// TIA Portal project "Catalyst_syzygy_v2.1" (V17) (continued)
VERSION : 0.1
   VAR
      ConnectP : TCON_IP_v4;
      MBControl : Struct
         diconnect : Bool;
      END_STRUCT;
   END_VAR
BEGIN
   ConnectP.InterfaceId := 258;
   ConnectP.ID := 16#1;
   ConnectP.ConnectionType := 11;
   ConnectP.LocalPort := 502;
END_DATA_BLOCK

DATA_BLOCK "TC-402B_DB"   // DB425
{ S7_Optimized_Access := 'TRUE' }
VERSION : 0.1
   VAR
      Data : "EurothermCtls_UDT";
      AddrCtrl : Struct
         CurrentAddr : UDInt;
         Down : Bool;
         Up : Bool;
         RisingUp : Bool;
      END_STRUCT;
   END_VAR
BEGIN
END_DATA_BLOCK

DATA_BLOCK "TC-402B_R1"   // DB429
{ S7_Optimized_Access := 'TRUE' }
AUTHOR : JL
VERSION : 0.1
// stored: InstanceOfName Eurotherm_MB_FB
"Eurotherm_MB_FB"
BEGIN
END_DATA_BLOCK

DATA_BLOCK "TC-402B_R2"   // DB431
{ S7_Optimized_Access := 'TRUE' }
AUTHOR : JL
VERSION : 0.1
// stored: InstanceOfName Eurotherm_MB_FB
"Eurotherm_MB_FB"
BEGIN
END_DATA_BLOCK

DATA_BLOCK "TC-402B_R3"   // DB432
{ S7_Optimized_Access := 'TRUE' }
AUTHOR : JL
VERSION : 0.1
// stored: InstanceOfName Eurotherm_MB_FB
"Eurotherm_MB_FB"
BEGIN
END_DATA_BLOCK

DATA_BLOCK "TC-402B_W1"   // DB435
{ S7_Optimized_Access := 'TRUE' }
AUTHOR : JL
VERSION : 0.1
// stored: InstanceOfName Eurotherm_MB_FB
"Eurotherm_MB_FB"
BEGIN
END_DATA_BLOCK

// folder: Outside Comms/ModBus Comms/MFCs/MFC-4011

DATA_BLOCK "MFC-4011_MB_R_DB"   // DB93
{ S7_Optimized_Access := 'TRUE' }
VERSION : 0.1
// stored: InstanceOfName MFC_MB_rDT
"MFC_MB_rDT"
BEGIN
END_DATA_BLOCK

DATA_BLOCK "MFC-4011_MB_W_DB"   // DB130
{ S7_Optimized_Access := 'TRUE' }
VERSION : 0.1
// stored: InstanceOfName MFC_MB_rDT
"MFC_MB_rDT"
BEGIN
END_DATA_BLOCK

DATA_BLOCK "MFC-4011_MB_RCMD_DB"   // DB133
{ S7_Optimized_Access := 'TRUE' }
AUTHOR : JL
VERSION : 0.1
// stored: InstanceOfName MFC_MB_iDT
"MFC_MB_iDT"
BEGIN
END_DATA_BLOCK

DATA_BLOCK "MFC-4011_MB_WCMD_DB"   // DB139
{ S7_Optimized_Access := 'TRUE' }
AUTHOR : JL
VERSION : 0.1
// stored: InstanceOfName MFC_MB_iDT
"MFC_MB_iDT"
BEGIN
END_DATA_BLOCK

DATA_BLOCK "MFC-4011_DB_MB"   // DB144
TITLE = MFC-4011 Modbus DB
{ S7_Optimized_Access := 'TRUE' }
VERSION : 0.1
   VAR
      Data : "AlicatCtl_UDT";
   END_VAR
BEGIN
END_DATA_BLOCK

// folder: Outside Comms/ModBus Comms/MFCs/MFC-4012

DATA_BLOCK "MFC-4012_MB_R_DB"   // DB200
{ S7_Optimized_Access := 'TRUE' }
VERSION : 0.1
// stored: InstanceOfName MFC_MB_rDT
"MFC_MB_rDT"
BEGIN
END_DATA_BLOCK

DATA_BLOCK "MFC-4012_MB_W_DB"   // DB201
{ S7_Optimized_Access := 'TRUE' }
VERSION : 0.1
// stored: InstanceOfName MFC_MB_rDT
"MFC_MB_rDT"
BEGIN
END_DATA_BLOCK

DATA_BLOCK "MFC-4012_MB_RCMD_DB"   // DB202
{ S7_Optimized_Access := 'TRUE' }
AUTHOR : JL
VERSION : 0.1
// stored: InstanceOfName MFC_MB_iDT
"MFC_MB_iDT"
BEGIN
END_DATA_BLOCK

DATA_BLOCK "MFC-4012_MB_WCMD_DB"   // DB239
{ S7_Optimized_Access := 'TRUE' }
AUTHOR : JL
VERSION : 0.1
// stored: InstanceOfName MFC_MB_iDT
"MFC_MB_iDT"
BEGIN
END_DATA_BLOCK

DATA_BLOCK "MFC-4012_DB_MB"   // DB240
TITLE = MFC-4011 Modbus DB
{ S7_Optimized_Access := 'TRUE' }
VERSION : 0.1
   VAR
      Data : "AlicatCtl_UDT";
   END_VAR
BEGIN
END_DATA_BLOCK

// folder: Outside Comms/ModBus Comms/MFCs/MFC-4021

DATA_BLOCK "MFC-4021_MB_R_DB"   // DB421
{ S7_Optimized_Access := 'TRUE' }
VERSION : 0.1
// stored: InstanceOfName MFC_MB_rDT
"MFC_MB_rDT"
BEGIN
END_DATA_BLOCK

DATA_BLOCK "MFC-4021_MB_W_DB"   // DB422
{ S7_Optimized_Access := 'TRUE' }
VERSION : 0.1
// stored: InstanceOfName MFC_MB_rDT
"MFC_MB_rDT"
BEGIN
END_DATA_BLOCK

DATA_BLOCK "MFC-4021_MB_RCMD_DB"   // DB423
{ S7_Optimized_Access := 'TRUE' }
AUTHOR : JL
VERSION : 0.1
// stored: InstanceOfName MFC_MB_iDT
"MFC_MB_iDT"
BEGIN
END_DATA_BLOCK

DATA_BLOCK "MFC-4021_MB_WCMD_DB"   // DB426
{ S7_Optimized_Access := 'TRUE' }
AUTHOR : JL
VERSION : 0.1
// stored: InstanceOfName MFC_MB_iDT
"MFC_MB_iDT"
BEGIN
END_DATA_BLOCK

DATA_BLOCK "MFC-4021_DB_MB"   // DB427
TITLE = MFC-4011 Modbus DB
{ S7_Optimized_Access := 'TRUE' }
VERSION : 0.1
   VAR
      Data : "AlicatCtl_UDT";
   END_VAR
BEGIN
END_DATA_BLOCK

// folder: Outside Comms/ModBus Comms/MFCs/MFC-4024

DATA_BLOCK "MFC-4024_MB_R_DB"   // DB388
{ S7_Optimized_Access := 'TRUE' }
VERSION : 0.1
// stored: InstanceOfName MFC_MB_rDT
"MFC_MB_rDT"
BEGIN
END_DATA_BLOCK

DATA_BLOCK "MFC-4024_MB_W_DB"   // DB390
{ S7_Optimized_Access := 'TRUE' }
VERSION : 0.1
// stored: InstanceOfName MFC_MB_rDT
"MFC_MB_rDT"
BEGIN
END_DATA_BLOCK

DATA_BLOCK "MFC-4024_MB_RCMD_DB"   // DB393
{ S7_Optimized_Access := 'TRUE' }
AUTHOR : JL
VERSION : 0.1
// stored: InstanceOfName MFC_MB_iDT
"MFC_MB_iDT"
BEGIN
END_DATA_BLOCK

DATA_BLOCK "MFC-4024_MB_WCMD_DB"   // DB395
{ S7_Optimized_Access := 'TRUE' }
AUTHOR : JL
VERSION : 0.1
// stored: InstanceOfName MFC_MB_iDT
"MFC_MB_iDT"
BEGIN
END_DATA_BLOCK

DATA_BLOCK "MFC-4024_DB_MB"   // DB396
TITLE = MFC-4011 Modbus DB
{ S7_Optimized_Access := 'TRUE' }
VERSION : 0.1
   VAR
      Data : "AlicatCtl_UDT";
   END_VAR
BEGIN
END_DATA_BLOCK

// folder: Outside Comms/ModBus Comms/MFCs/MFC-4025

DATA_BLOCK "MFC-4025_MB_R_DB"   // DB389
{ S7_Optimized_Access := 'TRUE' }
VERSION : 0.1
// stored: InstanceOfName MFC_MB_rDT
"MFC_MB_rDT"
BEGIN
END_DATA_BLOCK

DATA_BLOCK "MFC-4025_MB_W_DB"   // DB391
{ S7_Optimized_Access := 'TRUE' }
VERSION : 0.1
// stored: InstanceOfName MFC_MB_rDT
"MFC_MB_rDT"
BEGIN
END_DATA_BLOCK

DATA_BLOCK "MFC-4025_MB_RCMD_DB"   // DB392
{ S7_Optimized_Access := 'TRUE' }
AUTHOR : JL
VERSION : 0.1
// stored: InstanceOfName MFC_MB_iDT
"MFC_MB_iDT"
BEGIN
END_DATA_BLOCK

DATA_BLOCK "MFC-4025_MB_WCMD_DB"   // DB394
{ S7_Optimized_Access := 'TRUE' }
AUTHOR : JL
VERSION : 0.1
// stored: InstanceOfName MFC_MB_iDT
"MFC_MB_iDT"
BEGIN
END_DATA_BLOCK

DATA_BLOCK "MFC-4025_DB_MB"   // DB397
TITLE = MFC-4011 Modbus DB
{ S7_Optimized_Access := 'TRUE' }
VERSION : 0.1
   VAR
      Data : "AlicatCtl_UDT";
   END_VAR
BEGIN
END_DATA_BLOCK

// folder: Outside Comms/ModBus Comms/pH Transmitters/pH-2011/12

DATA_BLOCK "pH-2021_22_MB_rDT_DB"   // DB370
{ S7_Optimized_Access := 'TRUE' }
AUTHOR : JL
VERSION : 0.1
// stored: InstanceOfName MFC_MB_rDT
"MFC_MB_rDT"
BEGIN
END_DATA_BLOCK

DATA_BLOCK "pH-2011_12_MB_rDT_DB"   // DB371
{ S7_Optimized_Access := 'TRUE' }
AUTHOR : JL
VERSION : 0.1
// stored: InstanceOfName MFC_MB_rDT
"MFC_MB_rDT"
BEGIN
END_DATA_BLOCK

// folder: PID Controller/FlowControllers/DataBlocks

DATA_BLOCK "FIC-2011_DB"   // DB180
{ S7_Optimized_Access := 'TRUE' }
VERSION : 0.1
// stored: InstanceOfName PID_TIA
"PID_TIA"
BEGIN
   processVariableUpperLimit := 5.0;
   hmi.Config.P := 4.0;
   hmi.Config.I := 0.5;
END_DATA_BLOCK

DATA_BLOCK "FIC-2021_DB"   // DB182
{ S7_Optimized_Access := 'TRUE' }
VERSION : 0.1
// stored: InstanceOfName PID_TIA
"PID_TIA"
BEGIN
   processVariableUpperLimit := 5.0;
   hmi.Config.P := 4.0;
   hmi.Config.I := 0.5;
END_DATA_BLOCK

DATA_BLOCK "FIC-2012_DB"   // DB224
{ S7_Optimized_Access := 'TRUE' }
VERSION : 0.1
// stored: InstanceOfName PID_TIA
"PID_TIA"
BEGIN
   processVariableUpperLimit := 5.0;
   hmi.Config.P := 4.0;
   hmi.Config.I := 0.5;
END_DATA_BLOCK

DATA_BLOCK "FIC-2022_DB"   // DB225
{ S7_Optimized_Access := 'TRUE' }
VERSION : 0.1
// stored: InstanceOfName PID_TIA
"PID_TIA"
BEGIN
   processVariableUpperLimit := 5.0;
   hmi.Config.P := 4.0;
   hmi.Config.I := 0.5;
END_DATA_BLOCK

DATA_BLOCK "FIC-3011_DB"   // DB236
{ S7_Optimized_Access := 'TRUE' }
VERSION : 0.1
// stored: InstanceOfName PID_TIA
"PID_TIA"
BEGIN
   hmi.Config.P := 4.0;
   hmi.Config.I := 0.5;
END_DATA_BLOCK

// folder: PID Controller/Heater Controllers/DataBlocks

DATA_BLOCK "HFC-201_DB"   // DB150
{ S7_Optimized_Access := 'TRUE' }
VERSION : 0.1
// stored: InstanceOfName PID_TIA
"PID_TIA"
BEGIN
END_DATA_BLOCK

// folder: PID Controller/Level Controllers/DataBlocks

DATA_BLOCK "LIC-3011_DB"   // DB151
{ S7_Optimized_Access := 'TRUE' }
VERSION : 0.1
// stored: InstanceOfName PID_TIA
"PID_TIA"
BEGIN
END_DATA_BLOCK

// folder: PID Controller/PH Controllers/PHIC

DATA_BLOCK "PHIC-R-201_DB"   // DB132
{ S7_Optimized_Access := 'TRUE' }
VERSION : 0.1
// stored: InstanceOfName PID_TIA
"PID_TIA"
BEGIN
   hmi.Config.P := 5.0;
   hmi.Config.I := 4.0;
END_DATA_BLOCK

DATA_BLOCK "PHIC-R-202_DB"   // DB185
{ S7_Optimized_Access := 'TRUE' }
VERSION : 0.1
// stored: InstanceOfName PID_TIA
"PID_TIA"
BEGIN
   hmi.Config.P := 5.0;
   hmi.Config.I := 4.0;
END_DATA_BLOCK

// folder: PID Controller/PressureControllers

DATA_BLOCK "MFC-4012_DB"   // DB175
{ S7_Optimized_Access := 'TRUE' }
VERSION : 0.1
// stored: InstanceOfName PID_TIA
"PID_TIA"
BEGIN
   hmi.Config.P := 1.1;
   hmi.Config.I := 0.8;
END_DATA_BLOCK

// folder: PID Controller/PressureControllers/Datablocks

DATA_BLOCK "MFC-4011_DB"   // DB135
{ S7_Optimized_Access := 'TRUE' }
VERSION : 0.1
// stored: InstanceOfName PID_TIA
"PID_TIA"
BEGIN
   processVariableUpperLimit := 160.0;
   hmi.Config.P := 1.1;
   hmi.Config.I := 0.8;
END_DATA_BLOCK

DATA_BLOCK "MFC-4021_DB"   // DB136
{ S7_Optimized_Access := 'TRUE' }
VERSION : 0.1
// stored: InstanceOfName PID_TIA
"PID_TIA"
BEGIN
   processVariableUpperLimit := 160.0;
END_DATA_BLOCK

DATA_BLOCK "MFC-4025_DB"   // DB137
{ S7_Optimized_Access := 'TRUE' }
VERSION : 0.1
// stored: InstanceOfName PID_TIA
"PID_TIA"
BEGIN
   processVariableUpperLimit := 160.0;
END_DATA_BLOCK

DATA_BLOCK "MFC-4024_DB"   // DB138
{ S7_Optimized_Access := 'TRUE' }
VERSION : 0.1
// stored: InstanceOfName PID_TIA
"PID_TIA"
BEGIN
   processVariableUpperLimit := 160.0;
END_DATA_BLOCK

// folder: PID Controller/Temperature Controllers/DataBlocks

DATA_BLOCK "TIC-R402A_DB"   // DB149
{ S7_Optimized_Access := 'TRUE' }
VERSION : 0.1
// stored: InstanceOfName PID_TIA
"PID_TIA"
BEGIN
END_DATA_BLOCK

DATA_BLOCK "TIC-R402B_DB"   // DB154
{ S7_Optimized_Access := 'TRUE' }
VERSION : 0.1
// stored: InstanceOfName PID_TIA
"PID_TIA"
BEGIN
END_DATA_BLOCK

DATA_BLOCK "TIC-401_DB"   // DB160
{ S7_Optimized_Access := 'TRUE' }
VERSION : 0.1
// stored: InstanceOfName PID_TIA
"PID_TIA"
BEGIN
END_DATA_BLOCK

DATA_BLOCK "TIC-401_DB_1"   // DB188
{ S7_Optimized_Access := 'TRUE' }
VERSION : 0.1
// stored: InstanceOfName PID_TIA
"PID_TIA"
BEGIN
END_DATA_BLOCK

// folder: Pumps/Datablock

DATA_BLOCK "P-101A_DB"   // DB11
{ S7_Optimized_Access := 'TRUE' }
VERSION : 0.1
// stored: InstanceOfName SimpleMotorStater
"SimpleMotorStater"
BEGIN
END_DATA_BLOCK

DATA_BLOCK "P-101B_DB"   // DB17
{ S7_Optimized_Access := 'TRUE' }
VERSION : 0.1
// stored: InstanceOfName SimpleMotorStater
"SimpleMotorStater"
BEGIN
END_DATA_BLOCK

DATA_BLOCK "P-104A_DB"   // DB86
{ S7_Optimized_Access := 'TRUE' }
VERSION : 0.1
// stored: InstanceOfName SimpleMotorStater
"SimpleMotorStater"
BEGIN
   IL := true;
END_DATA_BLOCK

DATA_BLOCK "P-104B_DB"   // DB87
{ S7_Optimized_Access := 'TRUE' }
VERSION : 0.1
// stored: InstanceOfName SimpleMotorStater
"SimpleMotorStater"
BEGIN
   IL := true;
END_DATA_BLOCK

DATA_BLOCK "P-103A_DB"   // DB94
{ S7_Optimized_Access := 'TRUE' }
VERSION : 0.1
// stored: InstanceOfName SimpleMotorStater
"SimpleMotorStater"
BEGIN
END_DATA_BLOCK

DATA_BLOCK "P-201A_DB"   // DB95
{ S7_Optimized_Access := 'TRUE' }
VERSION : 0.1
// stored: InstanceOfName SimpleMotorStater
"SimpleMotorStater"
BEGIN
END_DATA_BLOCK

DATA_BLOCK "P-202A_DB"   // DB96
{ S7_Optimized_Access := 'TRUE' }
VERSION : 0.1
// stored: InstanceOfName SimpleMotorStater
"SimpleMotorStater"
BEGIN
END_DATA_BLOCK

DATA_BLOCK "P-301A_DB"   // DB97
{ S7_Optimized_Access := 'TRUE' }
VERSION : 0.1
// stored: InstanceOfName SimpleMotorStater
"SimpleMotorStater"
BEGIN
END_DATA_BLOCK

DATA_BLOCK "P-102A_DB"   // DB98
{ S7_Optimized_Access := 'TRUE' }
VERSION : 0.1
// stored: InstanceOfName SimpleMotorStater
"SimpleMotorStater"
BEGIN
END_DATA_BLOCK

DATA_BLOCK "P-102B_DB"   // DB100
{ S7_Optimized_Access := 'TRUE' }
VERSION : 0.1
// stored: InstanceOfName SimpleMotorStater
"SimpleMotorStater"
BEGIN
END_DATA_BLOCK

DATA_BLOCK "P-202B_DB"   // DB101
{ S7_Optimized_Access := 'TRUE' }
VERSION : 0.1
// stored: InstanceOfName SimpleMotorStater
"SimpleMotorStater"
BEGIN
END_DATA_BLOCK

DATA_BLOCK "P-103B_DB"   // DB102
{ S7_Optimized_Access := 'TRUE' }
VERSION : 0.1
// stored: InstanceOfName SimpleMotorStater
"SimpleMotorStater"
BEGIN
END_DATA_BLOCK

DATA_BLOCK "P-201B_DB"   // DB103
{ S7_Optimized_Access := 'TRUE' }
VERSION : 0.1
// stored: InstanceOfName SimpleMotorStater
"SimpleMotorStater"
BEGIN
END_DATA_BLOCK

DATA_BLOCK "P-301B_DB"   // DB105
{ S7_Optimized_Access := 'TRUE' }
VERSION : 0.1
// stored: InstanceOfName SimpleMotorStater
"SimpleMotorStater"
BEGIN
END_DATA_BLOCK

DATA_BLOCK "P-104C_DB"   // DB131
{ S7_Optimized_Access := 'TRUE' }
VERSION : 0.1
// stored: InstanceOfName SimpleMotorStater
"SimpleMotorStater"
BEGIN
END_DATA_BLOCK

// folder: Signal Inputs/LSHH

DATA_BLOCK "LSHH-1011_DB"   // DB76
{ S7_Optimized_Access := 'TRUE' }
VERSION : 1.1
// stored: InstanceOfName Signal
"Signal"
BEGIN
END_DATA_BLOCK

DATA_BLOCK "LSHH-1021_DB"   // DB77
{ S7_Optimized_Access := 'TRUE' }
VERSION : 1.1
// stored: InstanceOfName Signal
"Signal"
BEGIN
END_DATA_BLOCK

DATA_BLOCK "LSHH-1031_DB"   // DB78
{ S7_Optimized_Access := 'TRUE' }
VERSION : 1.1
// stored: InstanceOfName Signal
"Signal"
BEGIN
END_DATA_BLOCK

DATA_BLOCK "LSHH-2011_DB"   // DB79
{ S7_Optimized_Access := 'TRUE' }
VERSION : 1.1
// stored: InstanceOfName Signal
"Signal"
BEGIN
END_DATA_BLOCK

DATA_BLOCK "LSHH-2021_DB"   // DB156
{ S7_Optimized_Access := 'TRUE' }
VERSION : 1.1
// stored: InstanceOfName Signal
"Signal"
BEGIN
END_DATA_BLOCK

DATA_BLOCK "LSHH-1061_DB"   // DB237
{ S7_Optimized_Access := 'TRUE' }
VERSION : 1.1
// stored: InstanceOfName Signal
"Signal"
BEGIN
END_DATA_BLOCK

DATA_BLOCK "LSHH-1051_DB"   // DB238
{ S7_Optimized_Access := 'TRUE' }
VERSION : 1.1
// stored: InstanceOfName Signal
"Signal"
BEGIN
   Invert := true;
END_DATA_BLOCK

// folder: State MACHINE/1)Tanks/Tank T-101 (X)

DATA_BLOCK "T-101_DB"   // DB301
{ S7_Optimized_Access := 'TRUE' }
VERSION : 0.1
   VAR
      ExchangeCmds : Struct
         Send : Struct
            StartTank : Bool;
            ReqWater : Bool;
            StopReqWater : Bool;
            Release : Bool;
            Abort : Bool;
         END_STRUCT;
         Receive : Struct
            TankStarted : Bool;
            TankReady : Bool;
            PumpingOut : Bool;
            PumpsOff : Bool;
            Aborting : Bool;
         END_STRUCT;
      END_STRUCT;
      Cmds : "UnitCmds";
      Status : Struct
         Initializing : Bool;
         Ready : Bool;
         Running : Bool;
         PouringRunning : Bool;
         TankWashRunning : Bool;
         TubeWashRunning : Bool;
         Aborting : Bool;
         Status : Int;   // 1=Idle, 2=Running, 3=Stopping, 4=Held, 5=Holding
         "Step" : Int;
         State : Int;
      END_STRUCT;
      OS : Struct
         bit : Array[0..15] of Bool;   // One Shot Bit
      END_STRUCT;
      Equipments : Struct
         Valves : Struct
            "XV-1011" : "Cmd";
            "XV-1041" : "Cmd";
            "XV-1013" : "Cmd";
         END_STRUCT;
         Pumps : Struct
            "P-101A" : "Cmd";
            "P-101B" : "Cmd";
         END_STRUCT;
         VFD : Struct
            "VFD-1011" : "Cmd";
         END_STRUCT;
      END_STRUCT;
      PmpSel : Struct   // Pump Selection
         "P-101AB" : Int := 1;   // 1=P-101A, 2=P-101B
      END_STRUCT;
   END_VAR
BEGIN
END_DATA_BLOCK

DATA_BLOCK "T-101_Aux_DB"   // DB352
{ S7_Optimized_Access := 'TRUE' }
VERSION : 0.1
   VAR
      "Real" : Struct
         "FT-1041" : Struct
            SP : Real;
         END_STRUCT;
      END_STRUCT;
      "Timer" : Struct
         MinMixTimer : IEC_TIMER;
         PreMix : IEC_TIMER;   // Timer Premix
         "XV-1011" : IEC_TIMER;
         "XV-1041" : IEC_TIMER;
         "XV-1013" : IEC_TIMER;
      END_STRUCT;
      "Bool" : Struct
         MinMixT_Enab : Bool;
         MinMixT_Reset : Bool;
         PreMixTimer_Enab : Bool;   // Pre-Mix Timer Enable
         QtyWaterAdded : Bool;
         OperatorRequest : Bool;
         TOff : Bool;   // Turning Off Valves
      END_STRUCT;
      Constants : Struct
         CmdDelay : Time := T#2s;
      END_STRUCT;
   END_VAR
BEGIN
   "Timer".MinMixTimer.PT := T#30s;
END_DATA_BLOCK

DATA_BLOCK "T-101_SEQ_DB"   // DB357
{ S7_Optimized_Access := 'TRUE' }
VERSION : 0.1
// stored: InstanceOfName T-101_SEQ
"T-101_SEQ"
BEGIN
END_DATA_BLOCK

DATA_BLOCK "T-101_HMI_DB"   // DB360
{ S7_Optimized_Access := 'TRUE' }
VERSION : 0.1
   VAR
      FromHMI : "FromHMI";
      ToHMI : "ToHMI";
   END_VAR
BEGIN
   FromHMI.Procedure := 1;
END_DATA_BLOCK

// folder: State MACHINE/1)Tanks/Tank T-101 (X)/T-101 <---> R-201

DATA_BLOCK "T-101_Write_TO_R-201_DB"   // DB308
TITLE = Signal Exchange between R-201<->Reactor_Selector
{ S7_Optimized_Access := 'TRUE' }
VERSION : 0.1
   VAR
      TankStarted : Bool;   // Start Sequence
      Recirculating : Bool;
      PupmsOFF : Bool;   // Stop Sequence
      Abort : Bool;   // Abort Sequence
      RouteOpened : Bool;   // Transfer to Cooling Tank
      Idle : Bool;   // Held Sequence
   END_VAR
BEGIN
END_DATA_BLOCK

DATA_BLOCK "T-101_Read_FROM_R-201_DB"   // DB326
TITLE = Signal Exchange between R-201<->Reactor_Selector
{ S7_Optimized_Access := 'TRUE' }
VERSION : 0.1
   VAR
      StartPouring : Bool;
      ReactorStarted : Bool;
      OpenRoute : Bool;
      RouteOpened : Bool;
      Transfering : Bool;
      FillingDone : Bool;
      Aborting : Bool;
      Abort_Done : Bool;
      ReleaseTank : Bool;
      Idle : Bool;
   END_VAR
BEGIN
END_DATA_BLOCK

// folder: State MACHINE/1)Tanks/Tank T-101 (X)/T-101 <---> R-202

DATA_BLOCK "T-101_Write_TO_R-202_DB"   // DB292
TITLE = Signal Exchange between R-201<->Reactor_Selector
{ S7_Optimized_Access := 'TRUE' }
VERSION : 0.1
   VAR
      TankStarted : Bool;   // Start Sequence
      Recirculating : Bool;
      PupmsOFF : Bool;   // Stop Sequence
      Abort : Bool;   // Abort Sequence
      RouteOpened : Bool;   // Transfer to Cooling Tank
      Idle : Bool;   // Held Sequence
   END_VAR
BEGIN
END_DATA_BLOCK

DATA_BLOCK "T-101_Read_FROM_R-202_DB"   // DB322
TITLE = Signal Exchange between R-201<->Reactor_Selector
{ S7_Optimized_Access := 'TRUE' }
VERSION : 0.1
   VAR
      StartPouring : Bool;
      ReactorStarted : Bool;
      OpenRoute : Bool;
      RouteOpened : Bool;
      Transfering : Bool;
      FillingDone : Bool;
      Aborting : Bool;
      Abort_Done : Bool;
      ReleaseTank : Bool;
      Idle : Bool;
   END_VAR
BEGIN
END_DATA_BLOCK

// folder: State MACHINE/1)Tanks/Tank T-101 (X)/T-101 <---> T-104

DATA_BLOCK "T-101_Write_TO_T-104_DB"   // DB336
TITLE = Signal Exchange between R-201<->Reactor_Selector
{ S7_Optimized_Access := 'TRUE' }
VERSION : 0.1
   VAR
      StartTank : Bool;
      ReqWaterToWash : Bool;
      StopReqWaterToWash : Bool;
      ReqWaterToMix : Bool;
      StopReqWaterToMix : Bool;
      Release : Bool;
      Aborting : Bool;
      Abort_Done : Bool;
      Idle : Bool;
   END_VAR
BEGIN
END_DATA_BLOCK

DATA_BLOCK "T-101_Read_FROM_T-104_DB"   // DB340
TITLE = Signal Exchange between R-201<->Reactor_Selector
{ S7_Optimized_Access := 'TRUE' }
VERSION : 0.1
   VAR
      Wait : Bool;
      Started : Bool;   // Start Sequence
      Ready : Bool;
      Stop : Bool;   // Stop Sequence
      Abort : Bool;   // Abort Sequence
      Complete : Bool;
      Release : Bool;
      PARA : Bool;
      Initialization : Bool;
      PM : Bool;
      Monitoring : Bool;
      PumpingOut : Bool;   // Transfer to Cooling Tank
      PumpsOff : Bool;
      Held : Bool;   // Held Sequence
   END_VAR
BEGIN
END_DATA_BLOCK

// folder: State MACHINE/1)Tanks/Tank T-102 (Y)

DATA_BLOCK "T-102_DB"   // DB345
{ S7_Optimized_Access := 'TRUE' }
VERSION : 0.1
   VAR
      ExchangeCmds : Struct
         Send : Struct
            StartTank : Bool;
            ReqWater : Bool;
            StopReqWater : Bool;
            Release : Bool;
            Abort : Bool;
         END_STRUCT;
         Receive : Struct
            TankStarted : Bool;
            TankReady : Bool;
            PumpingOut : Bool;
            PumpsOff : Bool;
            Aborting : Bool;
         END_STRUCT;
      END_STRUCT;
      Cmds : "UnitCmds";
      Status : Struct
         Initializing : Bool;
         Ready : Bool;
         Running : Bool;
         PouringRunning : Bool;
         TankWashRunning : Bool;
         TubeWashRunning : Bool;
         Aborting : Bool;
         Status : Int;   // 1=Idle, 2=Running, 3=Stopping, 4=Held, 5=Holding
         "Step" : Int;
         State : Int;
      END_STRUCT;
      OS : Struct
         bit : Array[0..15] of Bool;   // One Shot Bit
      END_STRUCT;
      Equipments : Struct
         Valves : Struct
            "XV-1021" : "Cmd";
            "XV-1042" : "Cmd";
            "XV-1023" : "Cmd";
         END_STRUCT;
         Pumps : Struct
            "P-102A" : "Cmd";
            "P-102B" : "Cmd";
         END_STRUCT;
         VFD : Struct
            "VFD-1021" : "Cmd";
         END_STRUCT;
      END_STRUCT;
      PmpSel : Struct
         "P-102AB" : Int := 1;
      END_STRUCT;
   END_VAR
BEGIN
END_DATA_BLOCK

DATA_BLOCK "T-102_SEQ_DB"   // DB353
{ S7_Optimized_Access := 'TRUE' }
VERSION : 0.1
// stored: InstanceOfName T-102_SEQ
"T-102_SEQ"
BEGIN
END_DATA_BLOCK

DATA_BLOCK "T-102_HMI_DB"   // DB361
{ S7_Optimized_Access := 'TRUE' }
VERSION : 0.1
   VAR
      FromHMI : "FromHMI";
      ToHMI : "ToHMI";
   END_VAR
BEGIN
END_DATA_BLOCK

DATA_BLOCK "T-102_Aux_DB"   // DB364
{ S7_Optimized_Access := 'TRUE' }
VERSION : 0.1
   VAR
      "Real" : Struct
         "FT-1042" : Struct
            SP : Real;
         END_STRUCT;
      END_STRUCT;
      "Timer" : Struct
         MinMixTimer : IEC_TIMER;
         PreMix : IEC_TIMER;   // Timer Premix
         "XV-1021" : IEC_TIMER;
         "XV-1042" : IEC_TIMER;
         "XV-1023" : IEC_TIMER;
      END_STRUCT;
      "Bool" : Struct
         MinMixT_Enab : Bool;
         MinMixT_Reset : Bool;
         PreMixTimer_Enab : Bool;   // Pre-Mix Timer Enable
         QtyWaterAdded : Bool;
         OperatorRequest : Bool;
         TOff : Bool;   // Turning Off Valves
      END_STRUCT;
      Constants : Struct
         CmdDelay : Time := T#2s;
      END_STRUCT;
   END_VAR
BEGIN
   "Timer".MinMixTimer.PT := T#30s;
END_DATA_BLOCK

// folder: State MACHINE/1)Tanks/Tank T-102 (Y)/T-102 <---> R-201

DATA_BLOCK "T-102_Write_TO_R-201_DB"   // DB314
TITLE = Signal Exchange between R-201<->Reactor_Selector
{ S7_Optimized_Access := 'TRUE' }
VERSION : 0.1
   VAR
      TankStarted : Bool;   // Start Sequence
      Recirculating : Bool;
      PupmsOFF : Bool;   // Stop Sequence
      Abort : Bool;   // Abort Sequence
      RouteOpened : Bool;   // Transfer to Cooling Tank
      Idle : Bool;   // Held Sequence
   END_VAR
BEGIN
END_DATA_BLOCK

DATA_BLOCK "T-102_Read_FROM_R-201_DB"   // DB331
TITLE = Signal Exchange between R-201<->Reactor_Selector
{ S7_Optimized_Access := 'TRUE' }
VERSION : 0.1
   VAR
      StartPouring : Bool;
      ReactorStarted : Bool;
      OpenRoute : Bool;
      RouteOpened : Bool;
      Transfering : Bool;
      FillingDone : Bool;
      Aborting : Bool;
      Abort_Done : Bool;
      ReleaseTank : Bool;
      Idle : Bool;
   END_VAR
BEGIN
END_DATA_BLOCK

// folder: State MACHINE/1)Tanks/Tank T-102 (Y)/T-102 <---> R-202

DATA_BLOCK "T-102_Write_TO_R-202_DB"   // DB297
TITLE = Signal Exchange between R-201<->Reactor_Selector
{ S7_Optimized_Access := 'TRUE' }
VERSION : 0.1
   VAR
      TankStarted : Bool;   // Start Sequence
      Recirculating : Bool;
      PupmsOFF : Bool;   // Stop Sequence
      Abort : Bool;   // Abort Sequence
      RouteOpened : Bool;   // Transfer to Cooling Tank
      Idle : Bool;   // Held Sequence
   END_VAR
BEGIN
END_DATA_BLOCK

DATA_BLOCK "T-102_Read_FROM_R-202_DB"   // DB328
TITLE = Signal Exchange between R-201<->Reactor_Selector
{ S7_Optimized_Access := 'TRUE' }
VERSION : 0.1
   VAR
      StartPouring : Bool;
      ReactorStarted : Bool;
      OpenRoute : Bool;
      RouteOpened : Bool;
      Transfering : Bool;
      FillingDone : Bool;
      Aborting : Bool;
      Abort_Done : Bool;
      ReleaseTank : Bool;
      Idle : Bool;
   END_VAR
BEGIN
END_DATA_BLOCK

// folder: State MACHINE/1)Tanks/Tank T-102 (Y)/T-102 <---> T-104

DATA_BLOCK "T-102_Write_TO_T-104_DB"   // DB333
TITLE = Signal Exchange between R-201<->Reactor_Selector
{ S7_Optimized_Access := 'TRUE' }
VERSION : 0.1
   VAR
      StartTank : Bool;
      ReqWaterToWash : Bool;
      StopReqWaterToWash : Bool;
      ReqWaterToMix : Bool;
      StopReqWaterToMix : Bool;
      Release : Bool;
      Aborting : Bool;
      Abort_Done : Bool;
      Idle : Bool;
   END_VAR
BEGIN
END_DATA_BLOCK

DATA_BLOCK "T-102_Read_FROM_T-104_DB"   // DB342
TITLE = Signal Exchange between R-201<->Reactor_Selector
{ S7_Optimized_Access := 'TRUE' }
VERSION : 0.1
   VAR
      Wait : Bool;
      Started : Bool;   // Start Sequence
      Ready : Bool;
      Stop : Bool;   // Stop Sequence
      Abort : Bool;   // Abort Sequence
      Complete : Bool;
      Release : Bool;
      PARA : Bool;
      Initialization : Bool;
      PM : Bool;
      Monitoring : Bool;
      PumpingOut : Bool;   // Transfer to Cooling Tank
      PumpsOff : Bool;
      Held : Bool;   // Held Sequence
   END_VAR
BEGIN
END_DATA_BLOCK

// folder: State MACHINE/1)Tanks/Tank T-103 (Cooling Tank)

DATA_BLOCK "T-103_DB"   // DB272
{ S7_Optimized_Access := 'TRUE' }
VERSION : 0.1
   VAR
      ExchangeCmds : Struct
         Receive : Struct
            StartReceiving : Bool;   // Start from Reactors to Receive Material
            RequestProduct : Bool;   // Start from Centrifuge to send the Material
            OpenRoute : Bool;
            Transfering : Bool;
            TransferDone : Bool;
            Release : Bool;
            Idle : Bool;
         END_STRUCT;
         Send : Struct
            Started : Bool;
            RouteOpened : Bool;
            PumpingOut : Bool;
            PumpsOff : Bool;
            Release : Bool;
         END_STRUCT;
      END_STRUCT;
      Cmds : "UnitCmds";
      Tank : Struct
         Status : Int;   // 0= Ready to Receive, 1= Ready for Centerfuge
      END_STRUCT;
      Status : Struct
         Initializing : Bool;
         Ready : Bool;
         Running : Bool;
         Centrifuge : Bool;
         TankWashRunning : Bool;
         TubeWashRunning : Bool;
         Aborting : Bool;
         Status : Int;   // 1=Idle, 2=Running, 3=Stopping, 4=Held, 5=Holding
         "Step" : Int;
         State : Int;
      END_STRUCT;
      OS : Struct
         bit : Array[0..15] of Bool;   // One Shot Bit
      END_STRUCT;
      Equipments : Struct
         Valves : Struct
            "XV-1032" : "Cmd";
            "XV-1031" : "Cmd";
            "XV-3011" : "Cmd";
            "XV-1033" : "Cmd";
         END_STRUCT;
         Pumps : Struct
            "P-103A" : "Cmd";
            "P-103B" : "Cmd";
         END_STRUCT;
         VFD : Struct
            "VFD-T103" : "Cmd_VFD";
         END_STRUCT;
      END_STRUCT;
      PmpSel : Struct
         "P-103AB" : Int := 1;
      END_STRUCT;
   END_VAR
BEGIN
   Equipments.VFD."VFD-T103".p2000 := 1700.0;
END_DATA_BLOCK

DATA_BLOCK "T-103_SEQ_DB"   // DB274
{ S7_Optimized_Access := 'TRUE' }
VERSION : 0.1
// stored: InstanceOfName T-103_SEQ
"T-103_SEQ"
BEGIN
END_DATA_BLOCK

DATA_BLOCK "T-103_Aux_DB"   // DB355
{ S7_Optimized_Access := 'TRUE' }
VERSION : 0.1
   VAR
      "Real" : Struct
         "LT-1031" : Struct
            Min : Real;
         END_STRUCT;
      END_STRUCT;
      "Timer" : Struct
         StartRecircDelay : IEC_TIMER;
         "XV-1032" : IEC_TIMER;
         "XV-1031" : IEC_TIMER;
         "XV-3011" : IEC_TIMER;
         "XV-1033" : IEC_TIMER;
      END_STRUCT;
      "Bool" : Struct
         "VFD-T103" : Struct
            Start : Bool;
            Stop : Bool;
         END_STRUCT;
         StartRecirD_Enab : Bool;
         TOff : Bool;   // Turning Off Valves
      END_STRUCT;
      Constants : Struct
         CmdDelay : Time := T#2s;
      END_STRUCT;
   END_VAR
BEGIN
END_DATA_BLOCK

DATA_BLOCK "T-103_HMI_DB"   // DB362
{ S7_Optimized_Access := 'TRUE' }
VERSION : 0.1
   VAR
      FromHMI : "FromHMI";
      ToHMI : "ToHMI";
   END_VAR
BEGIN
END_DATA_BLOCK

// folder: State MACHINE/1)Tanks/Tank T-103 (Cooling Tank)/T-103 <---> Centrifuge

DATA_BLOCK "T-103_Write_TO_Centrifuge_DB"   // DB311
TITLE = Signal Exchange between R-201<->Reactor_Selector
{ S7_Optimized_Access := 'TRUE' }
VERSION : 0.1
   VAR
      Wait : Bool;
      ReadyToTranfer : Bool;   // Start Sequence
      Stop : Bool;   // Stop Sequence
      Abort : Bool;   // Abort Sequence
      Done : Bool;
      Release : Bool;
      PARA : Bool;
      Initialization : Bool;
      PM : Bool;
      Monitoring : Bool;
      RouteOpened : Bool;   // Transfer to Cooling Tank
      Transfering : Bool;
      Pumps_OFF : Bool;
      Idle : Bool;   // Held Sequence
   END_VAR
BEGIN
END_DATA_BLOCK

DATA_BLOCK "T-103_Read_FROM_Centrifuge_DB"   // DB321
TITLE = Signal Exchange between R-201<->Reactor_Selector
{ S7_Optimized_Access := 'TRUE' }
VERSION : 0.1
   VAR
      RequestProduct : Bool;   // Request Product
      OpenRoute : Bool;
      RouteOpened : Bool;
      "T-103_Empty" : Bool;
      BasketFull : Bool;   // Basket Full from Centrifuge
      FeelerRet : Bool;   // Feeler Retracted
      CloseRoute : Bool;
      Release : Bool;
   END_VAR
BEGIN
END_DATA_BLOCK

// folder: State MACHINE/1)Tanks/Tank T-103 (Cooling Tank)/T-103 <---> R-201

DATA_BLOCK "T-103_Write_TO_R-201_DB"   // DB284
TITLE = Signal Exchange between R-201<->Reactor_Selector
{ S7_Optimized_Access := 'TRUE' }
VERSION : 0.1
   VAR
      TankStarted : Bool;   // Start Sequence
      Stop : Bool;   // Stop Sequence
      Abort : Bool;   // Abort Sequence
      RouteOpened : Bool;   // Transfer to Cooling Tank
      ReleaseReactor : Bool;   // Release Reactor
      Held : Bool;   // Held Sequence
   END_VAR
BEGIN
END_DATA_BLOCK

DATA_BLOCK "T-103_Read_FROM_R-201_DB"   // DB291
TITLE = Signal Exchange between R-201<->Reactor_Selector
{ S7_Optimized_Access := 'TRUE' }
VERSION : 0.1
   VAR
      StartTank : Bool;
      OpenRoute : Bool;
      Transfering : Bool;
      TubWash_Done : Bool;
      Aborting : Bool;
      Abort_Done : Bool;
      "Transfer_To_T-103_Done" : Bool;
      Idle : Bool;
   END_VAR
BEGIN
END_DATA_BLOCK

// folder: State MACHINE/1)Tanks/Tank T-103 (Cooling Tank)/T-103 <--->R-202

DATA_BLOCK "T-103_Write_TO_R-202_DB"   // DB306
TITLE = Signal Exchange between R-201<->Reactor_Selector
{ S7_Optimized_Access := 'TRUE' }
VERSION : 0.1
   VAR
      TankStarted : Bool;   // Start Sequence
      Stop : Bool;   // Stop Sequence
      Abort : Bool;   // Abort Sequence
      RouteOpened : Bool;   // Transfer to Cooling Tank
      ReleaseReactor : Bool;   // Release Reactor
      Held : Bool;   // Held Sequence
   END_VAR
BEGIN
END_DATA_BLOCK

DATA_BLOCK "T-103_Read_FROM_R-202_DB"   // DB325
TITLE = Signal Exchange between R-201<->Reactor_Selector
{ S7_Optimized_Access := 'TRUE' }
VERSION : 0.1
   VAR
      StartTank : Bool;
      OpenRoute : Bool;
      Transfering : Bool;
      TubWash_Done : Bool;
      Abort_Done : Bool;
      "Transfer_To_T-103_Done" : Bool;
      Idle : Bool;
   END_VAR
BEGIN
END_DATA_BLOCK

// folder: State MACHINE/1)Tanks/Tank T-104 (Water System)

DATA_BLOCK "T-104_DB"   // DB302
{ S7_Optimized_Access := 'TRUE' }
VERSION : 0.1
   VAR
      ExchangeCmds : Struct
         Receive : Struct
            StartTank : Bool;
            ReqWater : Bool;
            StopReqWater : Bool;
            Release : Bool;
            Abort : Bool;
         END_STRUCT;
         Send : Struct
            TankStarted : Bool;
            TankReady : Bool;
            PumpingOut : Bool;
            PumpsOff : Bool;
            Aborting : Bool;
         END_STRUCT;
      END_STRUCT;
      Cmds : "UnitCmds";
      Status : Struct
         Initializing : Bool;
         Ready : Bool;
         Running : Bool;
         PouringRunning : Bool;
         TankWashRunning : Bool;
         TubeWashRunning : Bool;
         Aborting : Bool;
         Status : Int;   // 1=Idle, 2=Running, 3=Stopping, 4=Held, 5=Holding
         "Step" : Int;
         State : Int;
      END_STRUCT;
      OS : Struct
         bit : Array[0..15] of Bool;   // One Shot Bit
      END_STRUCT;
      Equipments : Struct
         "P-104A" : "Cmd";
         "P-104B" : "Cmd";
      END_STRUCT;
      PmpSel : Struct
         "P-104AB" : Int := 1;
      END_STRUCT;
   END_VAR
BEGIN
END_DATA_BLOCK

DATA_BLOCK "T-104_SEQ_DB"   // DB305
{ S7_Optimized_Access := 'TRUE' }
VERSION : 0.1
// stored: InstanceOfName T-104_SEQ
"T-104_SEQ"
BEGIN
END_DATA_BLOCK

DATA_BLOCK "T-104_HMI_DB"   // DB359
{ S7_Optimized_Access := 'TRUE' }
VERSION : 0.1
   VAR
      FromHMI : "FromHMI";
      ToHMI : "ToHMI";
   END_VAR
BEGIN
   FromHMI.Procedure := 1;
END_DATA_BLOCK

DATA_BLOCK "T-104_Aux_DB"   // DB369
{ S7_Optimized_Access := 'TRUE' }
VERSION : 0.1
   VAR
      "Real" : Struct
         "LT-xx" : Struct
            Min : Real;
         END_STRUCT;
      END_STRUCT;
      "Timer" : Struct
         xxxx : IEC_TIMER;
      END_STRUCT;
      "Bool" : Struct
         TOff : Bool;
      END_STRUCT;
   END_VAR
BEGIN
END_DATA_BLOCK

// folder: State MACHINE/1)Tanks/Tank T-104 (Water System)/T-104 <---> Centrifuge

